FUNCTION_BLOCK "FB_OptEthLink_V1.00"   // FB18, SCL
{ S7_Optimized_Access := 'TRUE' }
VERSION : 0.1
   VAR_INPUT
      IN_xCycleON : Bool;   // Cycle ON
      IN_xCycleONDel : Bool;   // Delayed cycle ON signal
      IN_xGeneralReset : Bool;   // General reset
      IN_xResetAlarms : Bool;   // Reset alarms
      IN_xFaultsEnabled : Bool;   // Faults enabled
      IN_tInterfaceID : Hw_Any;   // Interface ID
      IN_tSmallPckID : Conn_Ouc;   // Connection ID for small packets
      IN_tBigPckID : Conn_Ouc;   // Connection ID for big packets
      IN_uiSmallPckPort : UInt;   // Port small packet
      IN_uiBigPckPort : UInt;   // Port big packet
      IN_rgtStatusYCuts : Array[0.."DMAXYCUTBRIDGE_IND"] of Struct   // Status of YCut
         dDistanceSnapRoll_cmm : DInt;   // Distance from snaproll [mm/100]
         dBridgeStatus : DInt;   // Bridge actual status (1=OutOfProd 3=InProd 4=GlassBreak)
         rgxHeadProdOn : Array[0.."DMAXYHEADS_IND"] of Bool;   // Head#x production status
         rgxFireON : Array[0.."DMAXYHEADS_IND"] of Bool;   // Head#x fire status
         rgxArmON : Array[0.."DMAXYHEADS_IND"] of Bool;   // Head#x arm status
         rgdPosition_cmm : Array[0.."DMAXYHEADS_IND"] of DInt;   // Head#x position [mm/100]
      END_STRUCT;
      IN_rgtStatusXCuts : Array[0.."DMAXXHEADS_IND"] of Struct   // Status of XCuts
         dDistanceFromSnaproll_cmm : DInt;   // Distance from snaproll [mm/100]
         dStatus : DInt;   // XCut actual status (1=Idle 3=Running 7=Faulted)
         dActualCarriagePos_cmm : DInt;   // XCut actual carriage position [mm/100]
         dXCutActualStatus : DInt;   // XCut actual status (1=Disabled 3=Enabled)
         dCutTime_ms : DInt;   // XCut actual cutting time [ms]
      END_STRUCT;
      IN_rgtStatusMarker : Array[0..#DMAXMARKERS_IND] of Struct   // Status of Markers
         dHeadPosition_cmm : DInt;   // Actual head position [mm/100]
         dBridgeProdModeActual : DInt;   // Production modality actual (1=Out of production 3=In production 8=Out of production request 9=In production request)
         dDistanceFromSnaproll_cmm : DInt;   // Distance from snaproll [mm/100]
         dDistanceFromCenterLine_cmm : DInt;   // Distance from center line [mm/100]
         dSpraySpace_cmm : DInt;   // Spray space [mm/100]
         dSpare : DInt;
      END_STRUCT;
   END_VAR
   VAR_IN_OUT
      INO_tInitialize : "GP_OB_Initialize";   // Service bits
      INO_tEncoder : "UDT_Encoder";   // Encoder data
      INO_tOptimizer : "FB_OptManager_V1.00";   // Optimizer manager
      INO_tCaps : "UDT_CapData_Tracking";   // Cap data tracking
      INO_tDefects : "UDT_DefectData_Tracking_Ext";   // Defect data tracking
      INO_tMessage : "UDT_RP_TankMessages";   // Message tank
      INO_tAddMessageFromOpt : "UDT_RP_AddMessageCont_v2";   // Message add for received message
      INO_tAddMessageToOpt : "UDT_RP_AddMessageCont_v2";   // Message add for send message
      INO_xMessageAnomaly : Bool;   // Message anomaly bit
      INO_FB_Markers : "FB_Markers_V1.00";   // Markers FB
   END_VAR
   VAR
      AUX_tStatusPacket : Struct   // Status packet
         dTelID : DInt;   // Telegram identifier
         dTelCount : DInt;   // Telegram counter
         tServiceBit : Struct   // Services bits
            xSpare_24 : Bool;
            xSpare_25 : Bool;
            xSpare_26 : Bool;
            xSpare_27 : Bool;
            xSpare_28 : Bool;
            xSpare_29 : Bool;
            xSpare_30 : Bool;
            xSpare_31 : Bool;
            xSpare_16 : Bool;
            xSpare_17 : Bool;
            xSpare_18 : Bool;
            xSpare_19 : Bool;
            xSpare_20 : Bool;
            xSpare_21 : Bool;
            xSpare_22 : Bool;
            xSpare_23 : Bool;
            xOptRem : Bool;   // Optimizer in remote modality
            xGlassBreak : Bool;   // Glass break
            xSpare_10 : Bool;
            xSpare_11 : Bool;
            xSpare_12 : Bool;
            xSpare_13 : Bool;
            xSpare_14 : Bool;
            xSpare_15 : Bool;
            xSelPCA : Bool;   // Selection PC A
            xSelPCB : Bool;   // Selection PC B
            xSelPLCA : Bool;   // Selection PLC A
            xSelPLCB : Bool;   // Selection PLC B
            xSpare_4 : Bool;
            xSpare_5 : Bool;
            xSpare_6 : Bool;
            xSpare_7 : Bool;
         END_STRUCT;
         dActEnc_cmm : DInt;   // Actual encoder counter [mm/100]
         dActLehrSpeed_mm_min : DInt;   // Actuale lehr speed [mm/min]
         dDecLinePos_cmm : DInt;   // Decision line position [mm/100]
         dLastTargetEnc_cmm : DInt;   // Actual position last plate line [mm/100]
         dLastPlateID : DInt;   // Last plate ID
         dLastPlateLength_cmm : DInt;   // Last plate length [mm/100]
         dLastMapID : DInt;   // Last Map ID
         dSpare3 : DInt;   // Spare
         dRibbonGrossWidth_cmm : DInt;   // Ribbon gross width [mm/100]
         dSpare4 : DInt;   // Spare
         dRibbonNetWidth_cmm : DInt;   // Ribbon net width [mm/100]
         dRibbonWander_cmm : DInt;   // Ribbon wander [mm/100]
         dWanderRecTh_cmm : DInt;   // Ribbon wander recovery threshold [mm/100]
         dLineSpeed_mm_min : DInt;   // Line speed [mm/min]
         dSpare6 : DInt;   // Spare
         dSpare7 : DInt;   // Spare
         dSpare8 : DInt;   // Spare
         dSpare9 : DInt;   // Spare
         dSpare10 : DInt;   // Spare
         dSpare11 : DInt;   // Spare
         dBridgeAStatus : DInt;   // Bridge A status (1=OutOfProd 2=InProd 3=Locked)
         rgdBridgeAHeadxStatus : Array[0..#DMAXYHEADS_IND] of DInt;   // Bridge A headx status (1=OutOfProd 2=InProd 5=Firing)
         rgdBridgeAHeadPos_cmm : Array[0..#DMAXYHEADS_IND] of DInt;   // Bridge A headx position [mm/100]
         dSpare12 : DInt;
         dSpare13 : DInt;
         dSpare14 : DInt;
         dSpare15 : DInt;
         dSpare16 : DInt;
         dBridgeBStatus : DInt;   // Bridge B status (1=OutOfProd 2=InProd 3=Locked)
         rgdBridgeBHeadxStatus : Array[0..#DMAXYHEADS_IND] of DInt;   // Bridge B headx status (1=OutOfProd 2=InProd 5=Firing)
         rgdBridgeBHeadPos_cmm : Array[0..#DMAXYHEADS_IND] of DInt;   // Bridge B headx position [mm/100]
         rgdMarkerState : Array[0..#DMAXMARKERS_IND] of DInt;   // Markers state (1=OutOfProd 3=InProd 7=Anomaly)
         rgdMarkerPos_cmm : Array[0..#DMAXMARKERS_IND] of DInt;   // Markers actual position [mm/100]
         rgdMarkerDistSnap_cmm : Array[0..#DMAXMARKERS_IND] of DInt;   // Markers distance from snaproll [mm/100]
         rgdMarkerSprayTime_ms : Array[0..#DMAXMARKERS_IND] of DInt;   // Markers spray time [ms]
         rgdXCutsState : Array[0..#DMAXXCUT_IND] of DInt;   // XCuts state
         rgdXCutsTimes_ms : Array[0..#DMAXXCUT_IND] of DInt;   // XCuts timing [ms]
         dSpare22 : DInt;
      END_STRUCT;
      AUX_tPlatePacket : Struct   // Plate packet
         dTelID : DInt;   // Telegram identifier
         dTelCounter : DInt;   // Telegram counter
         dPlateHead_cmm : DInt;   // Plate head counter [mm/100]
         rgdLiteID : Array[0..#DMAXLITE_IND] of DInt;   // Lite ID
         rgdProductionID : Array[0..#DMAXLITE_IND] of DInt;   // Production ID
         rgdQualityID : Array[0..#DMAXLITE_IND] of DInt;   // Quality ID
         rgdLiteWidth_cmm : Array[0..#DMAXLITE_IND] of DInt;   // Lite width [mm/100]
         rgdDestMain : Array[0..#DMAXLITE_IND] of LInt;   // Main destination [mask]
         rgdDestAlt : Array[0..#DMAXLITE_IND] of LInt;   // Alternative destination [mask]
         rgdDest2Nd : Array[0..#DMAXLITE_IND] of LInt;   // Second choice destination [mask]
         rgdCulletCause : Array[0..#DMAXLITE_IND] of DInt;   // Cullet cause
         dNumLiteCap : DInt;   // Number of lites in cap
         dCapLength_cmm : DInt;   // Cap length [mm/100]
         dTotCapWidth_cmm : DInt;   // Total cap width [mm/100]
         dColorID : DInt;   // Color ID [mm/100]
         dCapThick_cmm : DInt;   // Cap thickness [mm/100]
         dGeomID : DInt;   // Geometrical ID
         dTrimWidthOper_cmm : DInt;   // Trim width operator side [mm/100]
         dTrimWidthOpOper_cmm : DInt;   // Trim width opposite operator side [mm/100]
         dWanderRec_cmm : DInt;   // Wander recoverd by YCut [mm/100]
         dYBridgeToCut : DInt;   // YCut bridge to cut
         rgxYHeadMask : Array[0..#DMAXYHEADSBITS_IND] of Bool;   // YCut head mask to cut
         rgYBridgePos_cmm : Array[0..#DMAXYHEADS_IND] of DInt;   // YCut head position
         rgxCutMissionHead : Array[0..#DMAXBITSXCUT_INDEX] of Bool;   // XCut mission head
         rgxCutMissionTail : Array[0..#DMAXBITSXCUT_INDEX] of Bool;   // XCut mission tail
         tGeneralFlags : Struct
            xClearCap : Bool;   // Clear cap
            xAutoTrim : Bool;   // Automatic trime selection
            xAutoSnap : Bool;   // Automatic snap bar selection
            xAutoSep : Bool;   // Automatic separator roll selection
            xTripleOpSide : Bool;   // Triple border on operator side
            xTripleOppoOpSide : Bool;   // Triple border on operator opposite side
            xDoubleBorder : Bool;   // Double border enabled
            xYCutSampleTest : Bool;   // YCut sample test
            xIsFixedCap : Bool;   // Is a fixed cap
            xSpare_9 : Bool;
            xSpare_10 : Bool;
            xSpare_11 : Bool;
            xSpare_12 : Bool;
            xSpare_13 : Bool;
            xSpare_14 : Bool;
            xSpare_15 : Bool;
            xSpare_16 : Bool;
            xSpare_17 : Bool;
            xSpare_18 : Bool;
            xSpare_19 : Bool;
            xSpare_20 : Bool;
            xSpare_21 : Bool;
            xSpare_22 : Bool;
            xSpare_23 : Bool;
            xSpare_24 : Bool;
            xSpare_25 : Bool;
            xSpare_26 : Bool;
            xSpare_27 : Bool;
            xSpare_28 : Bool;
            xSpare_29 : Bool;
            xSpare_30 : Bool;
            xSpare_31 : Bool;
         END_STRUCT;
         rgtLiteFlags : Array[0..#DMAXLITE_IND] of Struct
            xPow1Req : Bool;   // Powder #1 request
            xPow2Req : Bool;   // Powder #2 request
            xSatPlate : Bool;   // Saturation plate
            xGeomInsp : Bool;   // Geometrical inspection
            xPrint1 : Bool;   // Print #1 top
            xPrint2 : Bool;   // Print #1 bottom
            xSpare_6 : Bool;
            xSpare_7 : Bool;
            xSpare_8 : Bool;
            xSpare_9 : Bool;
            xSpare_10 : Bool;
            xSpare_11 : Bool;
            xSpare_12 : Bool;
            xSpare_13 : Bool;
            xSpare_14 : Bool;
            xSpare_15 : Bool;
            xMarkHomeHead : Bool;   // Laser mark home head
            xMarkHomeTail : Bool;   // Laser mark home tail
            xMarkCenterHead : Bool;   // Laser mark center head
            xMarkCenterTail : Bool;   // Laser mark center tail
            xMarkFarHead : Bool;   // Laser mark far head
            xMarkFarTail : Bool;   // Laser mark far tail
            xSpare_22 : Bool;
            xSpare_23 : Bool;
            xSpare_24 : Bool;
            xSpare_25 : Bool;
            xSpare_26 : Bool;
            xSpare_27 : Bool;
            xSpare_28 : Bool;
            xSpare_29 : Bool;
            xSpare_30 : Bool;
            xSpare_31 : Bool;   // This lite has a linked cap
         END_STRUCT;
         dExtBordOp : DInt;   // External border operator side
         dIntBordOp : DInt;   // Internal border operator side
         dExtBordOppoOp : DInt;   // External border opposite operator side
         dIntBordOppoOp : DInt;   // Internal border operator side
         rgdBumps : Array[0..#DMAXBUMP_IND] of DInt;   // Bumps splitter
         rgxChevrons : Array[0..#DMAXCHEVRON_IND] of Bool;   // Chevron rolls
         dPlateToPlate_cmm : DInt;   // Plate to plate distance [mm/100]
         dIndexPlateConv : DInt;   // Index plate convoy
         dMaxPlateConv : DInt;   // Max plate convoy
         dConvLength_cmm : DInt;   // Convoy length [mm/100]
         dMinWidth_cmm : DInt;   // Minimum width in production [mm/100]
         dMaxWidth_cmm : DInt;   // Maximum width in production [mm/100]
         dMinLength_cmm : DInt;   // Minimum length in production [mm/100]
         dMaxLength_cmm : DInt;   // Maximum length in production [mm/100]
         dCapID : DInt;   // Cap total ID
         rgdMapPlateID : Array[0..#DMAXLITE_IND] of DInt;   // Map plate ID
         dTripleEdgeOpSide_cmm : DInt;   // Triple edge operator side [mm/100]
         dTripleEdgeOppoOpSide_cmm : DInt;   // Triple edge operator opposite side [mm/100]
         dTripleEdgeHeadOpSide : DInt;   // Triple edge head selection operator side
         dTripleEdgeHeadOppoOpSide : DInt;   // Triple edge head selection oppositio operator side
         dFixedCapProdId : DInt;   // Fixed cap production ID
         rgdSpare : Array[0..10] of DInt;
      END_STRUCT;
      AUX_tDefectPacket : Struct   // Defect packet
         dTelID : DInt;   // Telegram identifier
         dTelCount : DInt;   // Telegram counter
         dNumDefect : DInt;   // Number of defect on packet
         dSpare : DInt;
         dSpare_1 : DInt;
         rgtDefects : Array[0..#DMAXDEFECTS_IND] of Struct
            dID : DInt;   // Defects ID
            dClass : DInt;   // Defects Class
            dSubtype : DInt;   // Defects Subtype
            dPosX_cmm : DInt;   // Defect position X [mm/100]
            dPosY_cmm : DInt;   // Defect position Y [mm/100]
            dTLength_cmm : DInt;   // Total length [mm/100]
            dTWidth_cmm : DInt;   // Total width [mm/100]
            dCLength_cmm : DInt;   // Core length [mm/100]
            dCWidth_cmm : DInt;   // Core width [mm/100]
            dDLength_cmm : DInt;   // Distortion length [mm/100]
            dDWidth_cmm : DInt;   // Distortion width [mm/100]
            dOptDist_mdptr : DInt;   // Optical distortion value [mdptr]
         END_STRUCT;
      END_STRUCT;
      AUX_tMessagePacketToOpt : Struct   // Message packet
         dTelID : DInt;   // Telegram identifier
         dTelCount : DInt;   // Telegram counter
         dNumMessage : DInt;   // Number of message on packet
         dSpare : DInt;
         rgtMessage : Array[0..#DMAXMESSAGEPACKET_IND] of Struct
            dCodeEvent : DInt;
            dEvent1 : DInt;
            dEvent2 : DInt;
            dEvent3 : DInt;
            dEvent4 : DInt;
            dEvent5 : DInt;
            dEvent6 : DInt;
            dEvent7 : DInt;
            dEvent8 : DInt;
            dEvent9 : DInt;
            dEvent10 : DInt;
         END_STRUCT;
      END_STRUCT;
      AUX_tMessagePacketFromOpt : Struct   // Message packet
         dTelID : DInt;   // Telegram identifier
         dTelCount : DInt;   // Telegram counter
         dNumMessage : DInt;   // Number of message on packet
         dSpare : DInt;
         rgtMessage : Array[0..#DMAXMESSAGEPACKET_IND] of Struct
            dCodeEvent : DInt;
            dEvent1 : DInt;
            dEvent2 : DInt;
            dEvent3 : DInt;
            dEvent4 : DInt;
            dEvent5 : DInt;
            dEvent6 : DInt;
            dEvent7 : DInt;
            dEvent8 : DInt;
            dEvent9 : DInt;
            dEvent10 : DInt;
         END_STRUCT;
      END_STRUCT;
      AUX_dNumPlatePacket : DInt;   // Number of plate on buffer
      AUX_rgtPlatePacketArray : Array[0..#DMAXPLATEPACKET_IND] of Struct   // Array buffer of plate
         dTelID : DInt;   // Telegram identifier
         dTelCounter : DInt;   // Telegram counter
         dPlateHead_cmm : DInt;   // Plate head counter [mm/100]
         rgdLiteID : Array[0..#DMAXLITE_IND] of DInt;   // Lite ID
         rgdProductionID : Array[0..#DMAXLITE_IND] of DInt;   // Production ID
         rgdQualityID : Array[0..#DMAXLITE_IND] of DInt;   // Quality ID
         rgdLiteWidth_cmm : Array[0..#DMAXLITE_IND] of DInt;   // Lite width [mm/100]
         rgdDestMain : Array[0..#DMAXLITE_IND] of LInt;   // Main destination [mask]
         rgdDestAlt : Array[0..#DMAXLITE_IND] of LInt;   // Alternative destination [mask]
         rgdDest2Nd : Array[0..#DMAXLITE_IND] of LInt;   // Second choice destination [mask]
         rgdCulletCause : Array[0..#DMAXLITE_IND] of DInt;   // Cullet cause
         dNumLiteCap : DInt;   // Number of lites in cap
         dCapLength_cmm : DInt;   // Cap length [mm/100]
         dTotCapWidth_cmm : DInt;   // Total cap width [mm/100]
         dColorID : DInt;   // Color ID [mm/100]
         dCapThick_cmm : DInt;   // Cap thickness [mm/100]
         dGeomID : DInt;   // Geometrical ID
         dTrimWidthOper_cmm : DInt;   // Trim width operator side [mm/100]
         dTrimWidthOpOper_cmm : DInt;   // Trim width opposite operator side [mm/100]
         dWanderRec_cmm : DInt;   // Wander recoverd by YCut [mm/100]
         dYBridgeToCut : DInt;   // YCut bridge to cut
         rgxYHeadMask : Array[0..#DMAXYHEADSBITS_IND] of Bool;   // YCut head mask to cut
         rgYBridgePos_cmm : Array[0..#DMAXYHEADS_IND] of DInt;   // YCut head position
         rgxCutMissionHead : Array[0..#DMAXBITSXCUT_INDEX] of Bool;   // XCut mission head
         rgxCutMissionTail : Array[0..#DMAXBITSXCUT_INDEX] of Bool;   // XCut mission tail
         tGeneralFlags : Struct
            xClearCap : Bool;   // Clear cap
            xAutoTrim : Bool;   // Automatic trime selection
            xAutoSnap : Bool;   // Automatic snap bar selection
            xAutoSep : Bool;   // Automatic separator roll selection
            xTripleOpSide : Bool;   // Triple border on operator side
            xTripleOppoOpSide : Bool;   // Triple border on operator opposite side
            xDoubleBorder : Bool;   // Double border enabled
            xYCutSampleTest : Bool;   // YCut sample test
            xIsFixedCap : Bool;   // Is a fixed cap
            xSpare_9 : Bool;
            xSpare_10 : Bool;
            xSpare_11 : Bool;
            xSpare_12 : Bool;
            xSpare_13 : Bool;
            xSpare_14 : Bool;
            xSpare_15 : Bool;
            xSpare_16 : Bool;
            xSpare_17 : Bool;
            xSpare_18 : Bool;
            xSpare_19 : Bool;
            xSpare_20 : Bool;
            xSpare_21 : Bool;
            xSpare_22 : Bool;
            xSpare_23 : Bool;
            xSpare_24 : Bool;
            xSpare_25 : Bool;
            xSpare_26 : Bool;
            xSpare_27 : Bool;
            xSpare_28 : Bool;
            xSpare_29 : Bool;
            xSpare_30 : Bool;
            xSpare_31 : Bool;
         END_STRUCT;
         rgtLiteFlags : Array[0..#DMAXLITE_IND] of Struct
            xPow1Req : Bool;   // Powder #1 request
            xPow2Req : Bool;   // Powder #2 request
            xSatPlate : Bool;   // Saturation plate
            xGeomInsp : Bool;   // Geometrical inspection
            xPrint1 : Bool;   // Print #1 top
            xPrint2 : Bool;   // Print #1 bottom
            xSpare_6 : Bool;
            xSpare_7 : Bool;
            xSpare_8 : Bool;
            xSpare_9 : Bool;
            xSpare_10 : Bool;
            xSpare_11 : Bool;
            xSpare_12 : Bool;
            xSpare_13 : Bool;
            xSpare_14 : Bool;
            xSpare_15 : Bool;
            xMarkHomeHead : Bool;   // Laser mark home head
            xMarkHomeTail : Bool;   // Laser mark home tail
            xMarkCenterHead : Bool;   // Laser mark center head
            xMarkCenterTail : Bool;   // Laser mark center tail
            xMarkFarHead : Bool;   // Laser mark far head
            xMarkFarTail : Bool;   // Laser mark far tail
            xSpare_22 : Bool;
            xSpare_23 : Bool;
            xSpare_24 : Bool;
            xSpare_25 : Bool;
            xSpare_26 : Bool;
            xSpare_27 : Bool;
            xSpare_28 : Bool;
            xSpare_29 : Bool;
            xSpare_30 : Bool;
            xSpare_31 : Bool;   // This lite has a linked cap
         END_STRUCT;
         dExtBordOp : DInt;   // External border operator side
         dIntBordOp : DInt;   // Internal border operator side
         dExtBordOppoOp : DInt;   // External border opposite operator side
         dIntBordOppoOp : DInt;   // Internal border operator side
         rgdBumps : Array[0..#DMAXBUMP_IND] of DInt;   // Bumps splitter
         rgxChevrons : Array[0..#DMAXCHEVRON_IND] of Bool;   // Chevron rolls
         dPlateToPlate_cmm : DInt;   // Plate to plate distance [mm/100]
         dIndexPlateConv : DInt;   // Index plate convoy
         dMaxPlateConv : DInt;   // Max plate convoy
         dConvLength_cmm : DInt;   // Convoy length [mm/100]
         dMinWidth_cmm : DInt;   // Minimum width in production [mm/100]
         dMaxWidth_cmm : DInt;   // Maximum width in production [mm/100]
         dMinLength_cmm : DInt;   // Minimum length in production [mm/100]
         dMaxLength_cmm : DInt;   // Maximum length in production [mm/100]
         dCapID : DInt;   // Cap total ID
         rgdMapPlateID : Array[0..#DMAXLITE_IND] of DInt;   // Map plate ID
         dTripleEdgeOpSide_cmm : DInt;   // Triple edge operator side [mm/100]
         dTripleEdgeOppoOpSide_cmm : DInt;   // Triple edge operator opposite side [mm/100]
         dTripleEdgeHeadOpSide : DInt;   // Triple edge head selection operator side
         dTripleEdgeHeadOppoOpSide : DInt;   // Triple edge head selection oppositio operator side
         dFixedCapProdId : DInt;   // Fixed cap production ID
         rgdSpare : Array[0..10] of DInt;
      END_STRUCT;
      AUX_rgb500SendBytePck : Array[0..#DSMALLSIZEPACKET_IND] of Byte;   // Byte array small size packet
      AUX_rgb500RecvBytePck : Array[0..#DSMALLSIZEPACKET_IND] of Byte;   // Byte array small size packet
      AUX_rgb1000SendBytePck : Array[0..#DBIGSIZEPACKET_IND] of Byte;   // Byte array big size packet
      AUX_rgb1000RecvBytePck : Array[0..#DBIGSIZEPACKET_IND] of Byte;   // Byte array big size packet
      FB_TSendSmall : TSEND_C;   // FB send small
      FB_TRecvSmall : TRCV_C;   // FB receive small
      FB_TSendBig : TSEND_C;   // FB send big
      FB_TRecvBig : TRCV_C;   // FB receive big
      AUX_tConnDataSmall : TCON_IP_v4;   // Connection small data structure
      AUX_tConnDataBig : TCON_IP_v4;   // Connection big data structure
      tPhasesNetworkSmall : Struct   // Phases network small
         xSendBuffer : Bool;   // Send buffer in progress
         xEndSendBuffer : Bool;   // End send buffer in progress
         xSpare2 : Bool;
         xSpare3 : Bool;
         xSpare4 : Bool;
         xSpare5 : Bool;
         xSpare6 : Bool;
         xSpare7 : Bool;
         xSpare8 : Bool;
         xSpare9 : Bool;
         xSpare10 : Bool;
         xSpare11 : Bool;
         xSpare12 : Bool;
         xSpare13 : Bool;
         xSpare14 : Bool;
         xSpare15 : Bool;
         xSpare16 : Bool;
         xSpare17 : Bool;
         xSpare18 : Bool;
         xSpare19 : Bool;
         xSpare20 : Bool;
         xSpare21 : Bool;
         xSpare22 : Bool;
         xSpare23 : Bool;
         xSpare24 : Bool;
         xSpare25 : Bool;
         xSpare26 : Bool;
         xSpare27 : Bool;
         xSpare28 : Bool;
         xSpare29 : Bool;
         xSpare30 : Bool;
         xSpare31 : Bool;
      END_STRUCT;
      tPhasesNetworkBig : Struct   // Phases network big
         xSendBuffer : Bool;   // Send buffer in progress
         xEndSendBuffer : Bool;   // End send buffer in progress
         xSpare2 : Bool;
         xSpare3 : Bool;
         xSpare4 : Bool;
         xSpare5 : Bool;
         xSpare6 : Bool;
         xSpare7 : Bool;
         xSpare8 : Bool;
         xSpare9 : Bool;
         xSpare10 : Bool;
         xSpare11 : Bool;
         xSpare12 : Bool;
         xSpare13 : Bool;
         xSpare14 : Bool;
         xSpare15 : Bool;
         xSpare16 : Bool;
         xSpare17 : Bool;
         xSpare18 : Bool;
         xSpare19 : Bool;
         xSpare20 : Bool;
         xSpare21 : Bool;
         xSpare22 : Bool;
         xSpare23 : Bool;
         xSpare24 : Bool;
         xSpare25 : Bool;
         xSpare26 : Bool;
         xSpare27 : Bool;
         xSpare28 : Bool;
         xSpare29 : Bool;
         xSpare30 : Bool;
         xSpare31 : Bool;
      END_STRUCT;
      AUX_xResetSendConnection : Bool;   // Reset send connection
      ST_xRetrySendTelegramSmall : Bool;   // Retry send telegram small
      ST_xRetrySendTelegramBig : Bool;   // Retry send telegram big
      ST_xStatusTelegramAvail : Bool;   // Status telegram available to send
      ST_xDefectTelegramAvail : Bool;   // Defect telegram available to send
      ST_xMessageTelegramAvail : Bool;   // Message telegram available to send
      ST_xSmallChannelConnected : Bool;   // Small channel connected
      ST_xBigChannelConnected : Bool;   // Big channel connected
      AUX_dWaitingNextStatus_ms : DInt;   // Waiting time for next status packet [ms]
   END_VAR
   VAR RETAIN
      AUX_dStatusTelegramCounter : DInt := 1;   // Status telegram counter
      AUX_dDefectTelegramCounter : DInt := 1;   // Defect telegram counter
      AUX_dMessageTelegramCounter : DInt := 1;   // Telegram message counter
   END_VAR
   VAR
      AUX_tEmptyMessage : "UDT_RP_Message_v2";   // Empty message
      tALM : Struct   // HMI Alarms
         tS : Struct   // Stopping faults
            xCh1NotCon : Bool;   // Channel 1 not connected {X|X|X|X|O}
            xCh2NotCon : Bool;   // Channel 2 not connected {X|X|X|X|O}
            xSpare_2 : Bool;
            xSpare_3 : Bool;
            xSpare_4 : Bool;
            xSpare_5 : Bool;
            xSpare_6 : Bool;
            xSpare_7 : Bool;
            xSpare_8 : Bool;
            xSpare_9 : Bool;
            xSpare_10 : Bool;
            xSpare_11 : Bool;
            xSpare_12 : Bool;
            xSpare_13 : Bool;
            xSpare_14 : Bool;
            xSpare_15 : Bool;
            xSpare_16 : Bool;
            xSpare_17 : Bool;
            xSpare_18 : Bool;
            xSpare_19 : Bool;
            xSpare_20 : Bool;
            xSpare_21 : Bool;
            xSpare_22 : Bool;
            xSpare_23 : Bool;
            xSpare_24 : Bool;
            xSpare_25 : Bool;
            xSpare_26 : Bool;
            xSpare_27 : Bool;
            xSpare_28 : Bool;
            xSpare_29 : Bool;
            xSpare_30 : Bool;
            xSpare_31 : Bool;
         END_STRUCT;
         tF : Struct   // Faults
            xSpare_0 : Bool;
            xSpare_1 : Bool;
            xSpare_2 : Bool;
            xSpare_3 : Bool;
            xSpare_4 : Bool;
            xSpare_5 : Bool;
            xSpare_6 : Bool;
            xSpare_7 : Bool;
            xSpare_8 : Bool;
            xSpare_9 : Bool;
            xSpare_10 : Bool;
            xSpare_11 : Bool;
            xSpare_12 : Bool;
            xSpare_13 : Bool;
            xSpare_14 : Bool;
            xSpare_15 : Bool;
            xSpare_16 : Bool;
            xSpare_17 : Bool;
            xSpare_18 : Bool;
            xSpare_19 : Bool;
            xSpare_20 : Bool;
            xSpare_21 : Bool;
            xSpare_22 : Bool;
            xSpare_23 : Bool;
            xSpare_24 : Bool;
            xSpare_25 : Bool;
            xSpare_26 : Bool;
            xSpare_27 : Bool;
            xSpare_28 : Bool;
            xSpare_29 : Bool;
            xSpare_30 : Bool;
            xSpare_31 : Bool;
         END_STRUCT;
         tW : Struct   // Warnings
            xSpare_0 : Bool;
            xSpare_1 : Bool;
            xSpare_2 : Bool;
            xSpare_3 : Bool;
            xSpare_4 : Bool;
            xSpare_5 : Bool;
            xSpare_6 : Bool;
            xSpare_7 : Bool;
            xSpare_8 : Bool;
            xSpare_9 : Bool;
            xSpare_10 : Bool;
            xSpare_11 : Bool;
            xSpare_12 : Bool;
            xSpare_13 : Bool;
            xSpare_14 : Bool;
            xSpare_15 : Bool;
            xSpare_16 : Bool;
            xSpare_17 : Bool;
            xSpare_18 : Bool;
            xSpare_19 : Bool;
            xSpare_20 : Bool;
            xSpare_21 : Bool;
            xSpare_22 : Bool;
            xSpare_23 : Bool;
            xSpare_24 : Bool;
            xSpare_25 : Bool;
            xSpare_26 : Bool;
            xSpare_27 : Bool;
            xSpare_28 : Bool;
            xSpare_29 : Bool;
            xSpare_30 : Bool;
            xSpare_31 : Bool;
         END_STRUCT;
      END_STRUCT;
   END_VAR
   VAR_TEMP
      TMP_dIndex : DInt;
      TMP_dSerializePos : DInt;   // Serialize temporary position
      TMP_iReturn : Int;
      TMP_dValue : DInt;
      TMP_dwMask : DWord;
      TMP_wMask : Word;
      TMP_dCounter : DInt;
      TMP_dRemaining : DInt;
      TMP_rgbDInt : Array[0..3] of Byte;
      TMP_iRetVal : Int;
      TMP_tNewMisMark : "UDT_Marker_Mission_Data";
      TMP_xCallAddTank : Bool;
      TMP_dwValue : DWord;
   END_VAR
   VAR CONSTANT
      DMAXYHEADS : DInt := 16;   // Maximum number of heads
      DMAXYHEADS_IND : DInt := 15;   // Maximum number of heads index (Always -1)
      DMAXYHEADSBITS : DInt := 32;   // Maximum number of heads bits
      DMAXYHEADSBITS_IND : DInt := 31;   // Maximum number of heads bits index (Always -1)
      DMAXMARKERS : DInt := 5;   // Maximum number of markers bridge
      DMAXMARKERS_IND : DInt := 4;   // Maximum number of markers bridge index (Always -1)
      DMAXXCUT : DInt := 5;   // Maximum number of cross cut bridge
      DMAXXCUT_IND : DInt := 4;   // Maximum number of cross cut bridge index (Always -1)
      DMAXLITE : DInt := 12;   // Maximum number of lite
      DMAXLITE_IND : DInt := 11;   // Maximum numer of lite index (Always -1)
      DMAXBITSXCUT : DInt := 32;   // Maximum number of request bits xcuts
      DMAXBITSXCUT_INDEX : DInt := 31;   // Maximum number of request bits xcuts index (Always -1)
      DMAXBUMP : DInt := 12;   // Maximum number of bump
      DMAXBUMP_IND : DInt := 11;   // Maximum numer of bump index (Always -1)
      DMAXCHEVRON : DInt := 32;   // Maximum number of chevron rolls
      DMAXCHEVRON_IND : DInt := 31;   // Maximum number of chevron rolls index (Always -1)
      BCONNTYPE : Byte := 16#0B;   // Optimizer connection type
      DSMALLSIZEPACKET : DInt := 500;   // Size of the small size packet
      DSMALLSIZEPACKET_IND : DInt := 499;   // Size of the small size packet index (Always -1)
      DBIGSIZEPACKET : DInt := 1000;   // Size of the big size packet
      DBIGSIZEPACKET_IND : DInt := 999;   // Size of the big size packet index (Always -1)
      DDELAYSTATUSPACKET_MS : DInt := 500;   // Status packet delay [ms]
      DSTATUSPACKETIDENT : DInt := 16#11111111;   // Status packet identifier
      DDEFECTPACKTIDENT : DInt := 16#22222222;   // Defect packet identifier
      DMESSAGEPACKETIDENT : DInt := 16#33333333;   // Message packet identifier
      DPLATEPACKTIDENT : DInt := 16#44444444;   // Plate packet identifier
      DMESSAGERECVPACKETIDENT : DInt := 16#55555555;   // Message received packet identifier
      DMAXTELEGRAMCOUNTER : DInt := 2000000000;   // Maximum telegram counter
      DMAXDEFECTS : DInt := 10;   // Maximum number of defects
      DMAXDEFECTS_IND : DInt := 9;   // Maximum number of defects index (Always -1)
      DMAXPLATEPACKET : DInt := 5;   // Number maximum of plate packet
      DMAXPLATEPACKET_IND : DInt := 4;   // Number maximum of plate packet index (Always -1)
      DMAXMESSAGEPACKET : DInt := 11;   // Number maximum of message packet
      DMAXMESSAGEPACKET_IND : DInt := 10;   // Number maximum of message packet index (Always -1)
   END_VAR
BEGIN
   IF #IN_xResetAlarms THEN

       #TMP_dwValue := 0;

       SCATTER(IN := #TMP_dwValue,
               OUT => #tALM.tS);

       SCATTER(IN := #TMP_dwValue,
               OUT => #tALM.tF);

       SCATTER(IN := #TMP_dwValue,
               OUT => #tALM.tW);


   END_IF;

   #ST_xSmallChannelConnected := TRUE;
   #ST_xBigChannelConnected := TRUE;

   IF #FB_TSendSmall.s_TDIAG_Status.State <> b#16#04(* OR #FB_TRecvSmall.s_TDIAG_Status.State <> b#16#04*) THEN

       #ST_xRetrySendTelegramSmall := FALSE;
       #ST_xStatusTelegramAvail := FALSE;
       #ST_xMessageTelegramAvail := FALSE;

       #tPhasesNetworkSmall.xSendBuffer := FALSE;
       #tPhasesNetworkSmall.xEndSendBuffer := FALSE;

       #ST_xSmallChannelConnected := FALSE;

       #INO_tDefects.xOptimizerRequireAllDef := TRUE;
   END_IF;

   IF #FB_TRecvBig.s_TRCV.ERROR  THEN
       #ST_xBigChannelConnected := FALSE;
   END_IF;

   //Calculate anomalies
   #tALM.tS.xCh1NotCon := NOT #ST_xSmallChannelConnected;
   #tALM.tS.xCh2NotCon := NOT #ST_xBigChannelConnected;


   IF #IN_xGeneralReset THEN
       #AUX_tConnDataSmall.InterfaceId := #IN_tInterfaceID;
       #AUX_tConnDataSmall.ID := #IN_tSmallPckID;
       #AUX_tConnDataSmall.ConnectionType := #BCONNTYPE;
       #AUX_tConnDataSmall.ActiveEstablished := FALSE;
       #AUX_tConnDataSmall.RemotePort := 0;
       #AUX_tConnDataSmall.LocalPort := #IN_uiSmallPckPort;

       #AUX_tConnDataBig.InterfaceId := #IN_tInterfaceID;
       #AUX_tConnDataBig.ID := #IN_tBigPckID;
       #AUX_tConnDataBig.ConnectionType := #BCONNTYPE;
       #AUX_tConnDataBig.ActiveEstablished := FALSE;
       #AUX_tConnDataBig.RemotePort := 0;
       #AUX_tConnDataBig.LocalPort := #IN_uiBigPckPort;
   END_IF;

   #AUX_dWaitingNextStatus_ms-= #INO_tInitialize.OUT_dExecutionTime_ms;

   IF #AUX_dWaitingNextStatus_ms < 0 THEN
       #AUX_dWaitingNextStatus_ms := 0;
   END_IF;


   IF NOT #ST_xMessageTelegramAvail AND #ST_xSmallChannelConnected THEN

       IF #INO_tMessage.dNumberOfMessage > 0 THEN
           #AUX_tMessagePacketToOpt.dTelID := #DMESSAGEPACKETIDENT;
           #AUX_tMessagePacketToOpt.dTelCount := #AUX_dMessageTelegramCounter;

           #TMP_dCounter := 0;

           WHILE (#TMP_dCounter < #DMAXMESSAGEPACKET) AND (#TMP_dCounter < #INO_tMessage.dNumberOfMessage) DO

               #AUX_tMessagePacketToOpt.rgtMessage[#TMP_dCounter].dCodeEvent := #INO_tMessage.rgtMessages[#TMP_dCounter].dCodeEvent;
               #AUX_tMessagePacketToOpt.rgtMessage[#TMP_dCounter].dEvent1 := #INO_tMessage.rgtMessages[#TMP_dCounter].dEvent1;
               #AUX_tMessagePacketToOpt.rgtMessage[#TMP_dCounter].dEvent2 := #INO_tMessage.rgtMessages[#TMP_dCounter].dEvent2;
               #AUX_tMessagePacketToOpt.rgtMessage[#TMP_dCounter].dEvent3 := #INO_tMessage.rgtMessages[#TMP_dCounter].dEvent3;
               #AUX_tMessagePacketToOpt.rgtMessage[#TMP_dCounter].dEvent4 := #INO_tMessage.rgtMessages[#TMP_dCounter].dEvent4;
               #AUX_tMessagePacketToOpt.rgtMessage[#TMP_dCounter].dEvent5 := #INO_tMessage.rgtMessages[#TMP_dCounter].dEvent5;
               #AUX_tMessagePacketToOpt.rgtMessage[#TMP_dCounter].dEvent6 := #INO_tMessage.rgtMessages[#TMP_dCounter].dEvent6;
               #AUX_tMessagePacketToOpt.rgtMessage[#TMP_dCounter].dEvent7 := #INO_tMessage.rgtMessages[#TMP_dCounter].dEvent7;
               #AUX_tMessagePacketToOpt.rgtMessage[#TMP_dCounter].dEvent8 := #INO_tMessage.rgtMessages[#TMP_dCounter].dEvent8;
               #AUX_tMessagePacketToOpt.rgtMessage[#TMP_dCounter].dEvent9 := #INO_tMessage.rgtMessages[#TMP_dCounter].dEvent9;
               #AUX_tMessagePacketToOpt.rgtMessage[#TMP_dCounter].dEvent10 := #INO_tMessage.rgtMessages[#TMP_dCounter].dEvent10;

               #INO_tMessage.rgtMessages[#TMP_dCounter] := #AUX_tEmptyMessage;

               #TMP_dCounter += 1;

           END_WHILE;

           //Clear the remaining packet
           FOR #TMP_dIndex := #TMP_dCounter TO #DMAXMESSAGEPACKET - 1 DO
               #AUX_tMessagePacketToOpt.rgtMessage[#TMP_dIndex].dCodeEvent := 0;
               #AUX_tMessagePacketToOpt.rgtMessage[#TMP_dIndex].dEvent1 := 0;
               #AUX_tMessagePacketToOpt.rgtMessage[#TMP_dIndex].dEvent2 := 0;
               #AUX_tMessagePacketToOpt.rgtMessage[#TMP_dIndex].dEvent3 := 0;
               #AUX_tMessagePacketToOpt.rgtMessage[#TMP_dIndex].dEvent4 := 0;
               #AUX_tMessagePacketToOpt.rgtMessage[#TMP_dIndex].dEvent5 := 0;
               #AUX_tMessagePacketToOpt.rgtMessage[#TMP_dIndex].dEvent6 := 0;
               #AUX_tMessagePacketToOpt.rgtMessage[#TMP_dIndex].dEvent7 := 0;
               #AUX_tMessagePacketToOpt.rgtMessage[#TMP_dIndex].dEvent8 := 0;
               #AUX_tMessagePacketToOpt.rgtMessage[#TMP_dIndex].dEvent9 := 0;
               #AUX_tMessagePacketToOpt.rgtMessage[#TMP_dIndex].dEvent10 := 0;
           END_FOR;

           #AUX_tMessagePacketToOpt.dNumMessage := #TMP_dCounter;
           #AUX_dMessageTelegramCounter+= 1;
           #ST_xMessageTelegramAvail := TRUE;
           #TMP_dRemaining := #INO_tMessage.dNumberOfMessage - #TMP_dCounter;

           IF #TMP_dRemaining > 0 THEN
               #TMP_iRetVal :=  MOVE_BLK_VARIANT(   SRC:= #INO_tMessage.rgtMessages, 
                                   COUNT:=DINT_TO_UDINT(#TMP_dRemaining), 
                                   SRC_INDEX:=#TMP_dCounter, 
                                   DEST_INDEX:=0, 
                                   DEST=>#INO_tMessage.rgtMessages);
               //Reset the remaining
               FOR #TMP_dIndex := #TMP_dRemaining TO #INO_tMessage.dNumberOfMessage - 1 DO
                   #INO_tMessage.rgtMessages[#TMP_dIndex] := #AUX_tEmptyMessage;
               END_FOR;

               #INO_tMessage.dNumberOfMessage := #TMP_dRemaining;

           ELSE
               #INO_tMessage.dNumberOfMessage := 0;
           END_IF;
       END_IF;
   END_IF;

   //Prepare defect telegram
   IF NOT #ST_xDefectTelegramAvail AND #ST_xSmallChannelConnected  THEN

       IF #INO_tDefects.tDefectsForOpt.dNumberOfDefect > 0 THEN

           #AUX_tDefectPacket.dTelID := #DDEFECTPACKTIDENT;
           #AUX_tDefectPacket.dTelCount := #AUX_dDefectTelegramCounter;
           #AUX_tDefectPacket.dNumDefect := #INO_tDefects.tDefectsForOpt.dNumberOfDefect;

           FOR #TMP_dIndex := 0 TO #DMAXDEFECTS_IND DO

               #AUX_tDefectPacket.rgtDefects[#TMP_dIndex].dID := #INO_tDefects.tDefectsForOpt.rgtDefects[#TMP_dIndex].dID;
               #AUX_tDefectPacket.rgtDefects[#TMP_dIndex].dClass := #INO_tDefects.tDefectsForOpt.rgtDefects[#TMP_dIndex].dClass;
               #AUX_tDefectPacket.rgtDefects[#TMP_dIndex].dSubtype := #INO_tDefects.tDefectsForOpt.rgtDefects[#TMP_dIndex].dSubType;
               #AUX_tDefectPacket.rgtDefects[#TMP_dIndex].dPosX_cmm := #INO_tDefects.tDefectsForOpt.rgtDefects[#TMP_dIndex].dXPosition_cmm;
               #AUX_tDefectPacket.rgtDefects[#TMP_dIndex].dPosY_cmm := #INO_tDefects.tDefectsForOpt.rgtDefects[#TMP_dIndex].dYPosition_cmm;
               #AUX_tDefectPacket.rgtDefects[#TMP_dIndex].dCLength_cmm := #INO_tDefects.tDefectsForOpt.rgtDefects[#TMP_dIndex].dCoreLength_um;
               #AUX_tDefectPacket.rgtDefects[#TMP_dIndex].dCWidth_cmm := #INO_tDefects.tDefectsForOpt.rgtDefects[#TMP_dIndex].dCoreWidth_um;
               #AUX_tDefectPacket.rgtDefects[#TMP_dIndex].dDLength_cmm := #INO_tDefects.tDefectsForOpt.rgtDefects[#TMP_dIndex].dDistLength_um;
               #AUX_tDefectPacket.rgtDefects[#TMP_dIndex].dDWidth_cmm := #INO_tDefects.tDefectsForOpt.rgtDefects[#TMP_dIndex].dDistWidth_um;
               #AUX_tDefectPacket.rgtDefects[#TMP_dIndex].dTLength_cmm := #INO_tDefects.tDefectsForOpt.rgtDefects[#TMP_dIndex].dTotalLength_um;
               #AUX_tDefectPacket.rgtDefects[#TMP_dIndex].dTWidth_cmm := #INO_tDefects.tDefectsForOpt.rgtDefects[#TMP_dIndex].dTotalWidth_um;
               #AUX_tDefectPacket.rgtDefects[#TMP_dIndex].dOptDist_mdptr := #INO_tDefects.tDefectsForOpt.rgtDefects[#TMP_dIndex].dOptValue_mdptr;

           END_FOR;

           #ST_xDefectTelegramAvail := TRUE;
           #AUX_dDefectTelegramCounter += 1;
           #INO_tDefects.tDefectsForOpt.dNumberOfDefect := 0;
       END_IF;

   END_IF;

   //Prepare status telegram
   IF NOT #ST_xStatusTelegramAvail AND #AUX_dWaitingNextStatus_ms = 0 AND #ST_xSmallChannelConnected THEN

       #AUX_dWaitingNextStatus_ms := #DDELAYSTATUSPACKET_MS;

       //Prepare data
       #AUX_tStatusPacket.dTelID :=  #DSTATUSPACKETIDENT;
       #AUX_tStatusPacket.dSpare22 := #DSTATUSPACKETIDENT;
       #AUX_tStatusPacket.dTelCount := #AUX_dStatusTelegramCounter;


       IF "FB_OptManager_V1_00_IDB".tHMR.dSelOptimizer = 1 THEN
           #AUX_tStatusPacket.tServiceBit.xSelPCA := TRUE;
           #AUX_tStatusPacket.tServiceBit.xSelPCB := FALSE;
       ELSE
           #AUX_tStatusPacket.tServiceBit.xSelPCA := FALSE;
           #AUX_tStatusPacket.tServiceBit.xSelPCB := TRUE;
       END_IF;

       #AUX_tStatusPacket.tServiceBit.xSelPLCA := TRUE;
       #AUX_tStatusPacket.tServiceBit.xSelPLCB := FALSE;
       #AUX_tStatusPacket.tServiceBit.xOptRem := TRUE;
       #AUX_tStatusPacket.tServiceBit.xGlassBreak := FALSE;

       #AUX_tStatusPacket.dActEnc_cmm := #INO_tEncoder.dActualEncoderCounter_cmm;
       #AUX_tStatusPacket.dActLehrSpeed_mm_min := #INO_tEncoder.dActSpeedValue_mm_min;
       #AUX_tStatusPacket.dDecLinePos_cmm := #INO_tOptimizer.tHMR.dDecisionLinePosition_cmm;
       #AUX_tStatusPacket.dLastTargetEnc_cmm := #INO_tCaps.dLastTargetLineValue_cmm;
       #AUX_tStatusPacket.dLastPlateID := #INO_tCaps.dLastValidCapID;

       #AUX_tStatusPacket.dRibbonGrossWidth_cmm := #INO_tOptimizer.tHMR.rgtRibbonData[#INO_tOptimizer.tHMW.dSelectRibbonDataSource].dGrossWidth_cmm;
       #AUX_tStatusPacket.dRibbonNetWidth_cmm := #INO_tOptimizer.tHMR.rgtRibbonData[#INO_tOptimizer.tHMW.dSelectRibbonDataSource].dNetWidth_cmm;

       #AUX_tStatusPacket.dWanderRecTh_cmm := #INO_tOptimizer.tHMW.dWanderRecThr_cmm;

       IF #INO_tOptimizer.tHMW.dSelectWanderMode = 0 THEN
           #AUX_tStatusPacket.dRibbonWander_cmm := #INO_tOptimizer.tHMR.rgtRibbonData[#INO_tOptimizer.tHMW.dSelectWanderDataSource].dNetWander_cmm + #INO_tOptimizer.tHMW.dWanderOffset_cmm;
       ELSE
           #AUX_tStatusPacket.dRibbonWander_cmm := #INO_tOptimizer.tHMR.rgtRibbonData[#INO_tOptimizer.tHMW.dSelectWanderDataSource].dGrossWander_cmm + #INO_tOptimizer.tHMW.dWanderOffset_cmm;
       END_IF;


       CASE #IN_rgtStatusYCuts[0].dBridgeStatus OF

           1:
               #AUX_tStatusPacket.dBridgeAStatus := 1;//Out of production
           3: #AUX_tStatusPacket.dBridgeAStatus := 2;
           4: #AUX_tStatusPacket.dBridgeAStatus := 2; //Glass break, out of production for optimizer

       END_CASE;

       CASE #IN_rgtStatusYCuts[1].dBridgeStatus OF

           1:
               #AUX_tStatusPacket.dBridgeBStatus := 1;//Out of production
           3: #AUX_tStatusPacket.dBridgeBStatus := 2;
           4: #AUX_tStatusPacket.dBridgeBStatus := 2; //Glass break, out of production for optimizer

       END_CASE;

       FOR #TMP_dIndex := 0 TO #DMAXYHEADS_IND DO

           IF #IN_rgtStatusYCuts[0].rgxHeadProdOn[#TMP_dIndex] = TRUE THEN
               #AUX_tStatusPacket.rgdBridgeAHeadxStatus[#TMP_dIndex] := 2;
           ELSE
               #AUX_tStatusPacket.rgdBridgeAHeadxStatus[#TMP_dIndex] := 1;
           END_IF;

           IF #IN_rgtStatusYCuts[1].rgxHeadProdOn[#TMP_dIndex] = TRUE THEN
               #AUX_tStatusPacket.rgdBridgeBHeadxStatus[#TMP_dIndex] := 2;
           ELSE
               #AUX_tStatusPacket.rgdBridgeBHeadxStatus[#TMP_dIndex] := 1;
           END_IF;

       END_FOR;

       #AUX_tStatusPacket.rgdBridgeAHeadPos_cmm := #IN_rgtStatusYCuts[0].rgdPosition_cmm;
       #AUX_tStatusPacket.rgdBridgeBHeadPos_cmm := #IN_rgtStatusYCuts[1].rgdPosition_cmm;

       FOR #TMP_dIndex := 0 TO #DMAXMARKERS_IND DO

           #AUX_tStatusPacket.rgdMarkerDistSnap_cmm[#TMP_dIndex] := #IN_rgtStatusMarker[#TMP_dIndex].dDistanceFromSnaproll_cmm;
           #AUX_tStatusPacket.rgdMarkerPos_cmm[#TMP_dIndex] := #IN_rgtStatusMarker[#TMP_dIndex].dHeadPosition_cmm;
           #AUX_tStatusPacket.rgdMarkerSprayTime_ms[#TMP_dIndex] := REAL_TO_DINT(DINT_TO_REAL(#IN_rgtStatusMarker[#TMP_dIndex].dSpraySpace_cmm) / #INO_tEncoder.rActSpeedValue_cmm_ms);

           CASE #IN_rgtStatusMarker[#TMP_dIndex].dBridgeProdModeActual OF

               1: #AUX_tStatusPacket.rgdMarkerState[#TMP_dIndex] := 1;//Out of production
               3: #AUX_tStatusPacket.rgdMarkerState[#TMP_dIndex] := 2;//In production
               8: #AUX_tStatusPacket.rgdMarkerState[#TMP_dIndex] := 1;//Out of production
               9: #AUX_tStatusPacket.rgdMarkerState[#TMP_dIndex] := 1;//Out of production

           END_CASE;

       END_FOR; 

       FOR #TMP_dIndex := 0 TO "DMAXXHEADS_IND" DO

           CASE #IN_rgtStatusXCuts[#TMP_dIndex].dXCutActualStatus OF

               1: #AUX_tStatusPacket.rgdXCutsState[#TMP_dIndex] := 0;
               3: #AUX_tStatusPacket.rgdXCutsState[#TMP_dIndex] := 1;

           END_CASE;

           #AUX_tStatusPacket.rgdXCutsTimes_ms[#TMP_dIndex] := #IN_rgtStatusXCuts[#TMP_dIndex].dCutTime_ms;

       END_FOR;

       IF #AUX_dStatusTelegramCounter >= #DMAXTELEGRAMCOUNTER THEN
           #AUX_dStatusTelegramCounter := 1;
       ELSE
           #AUX_dStatusTelegramCounter += 1;
       END_IF;

       #ST_xStatusTelegramAvail := TRUE;

   END_IF;


   #AUX_xResetSendConnection := #IN_xGeneralReset OR (#FB_TSendSmall.s_TDIAG_Status.State <> b#16#04 AND #IN_xResetAlarms);


   IF (NOT #tPhasesNetworkSmall.xEndSendBuffer) AND (NOT #tPhasesNetworkSmall.xSendBuffer) AND 
           ((#ST_xRetrySendTelegramSmall)OR (#ST_xStatusTelegramAvail)OR (#ST_xDefectTelegramAvail) OR (#ST_xMessageTelegramAvail)) THEN

       IF (NOT #ST_xRetrySendTelegramSmall) THEN

           IF (#ST_xStatusTelegramAvail) THEN
               #TMP_dSerializePos := 0;
               #TMP_iReturn := Serialize(SRC_VARIABLE:=#AUX_tStatusPacket, DEST_ARRAY=>#AUX_rgb500SendBytePck, POS:=#TMP_dSerializePos);    
               #ST_xStatusTelegramAvail := FALSE;
           ELSIF (#ST_xDefectTelegramAvail) THEN
               #TMP_dSerializePos := 0;
               #TMP_iReturn := Serialize(SRC_VARIABLE:=#AUX_tDefectPacket, DEST_ARRAY=>#AUX_rgb500SendBytePck, POS:=#TMP_dSerializePos);    
               #ST_xDefectTelegramAvail := FALSE;
           ELSIF (#ST_xMessageTelegramAvail) THEN
               #TMP_dSerializePos := 0;
               #TMP_iReturn := Serialize(SRC_VARIABLE:=#AUX_tMessagePacketToOpt, DEST_ARRAY=>#AUX_rgb500SendBytePck, POS:=#TMP_dSerializePos);    
               #ST_xMessageTelegramAvail := FALSE;
           END_IF;

       END_IF;

       #ST_xRetrySendTelegramSmall := FALSE;
       #tPhasesNetworkSmall.xSendBuffer := TRUE;

   END_IF;

   #FB_TRecvSmall(EN_R:=TRUE,
                CONT:=TRUE,
                CONNECT:=#AUX_tConnDataSmall,
                DATA:=#AUX_rgb500RecvBytePck,
                COM_RST:=#AUX_xResetSendConnection);

   #FB_TRecvBig(EN_R:=TRUE,
                CONT:=TRUE,
               LEN := 0,
                CONNECT:=#AUX_tConnDataBig,
                DATA:=#AUX_rgb1000RecvBytePck,
                COM_RST:=#AUX_xResetSendConnection);

   #FB_TSendSmall(REQ:=#tPhasesNetworkSmall.xSendBuffer,
             CONT:=TRUE,
             LEN:=0,
             CONNECT:=#AUX_tConnDataSmall,
             DATA:=#AUX_rgb500SendBytePck,
             COM_RST:=#AUX_xResetSendConnection);

   #FB_TSendBig(REQ:=#tPhasesNetworkBig.xSendBuffer,
             CONT:=TRUE,
             LEN:=0,
             CONNECT:=#AUX_tConnDataBig,
             DATA:=#AUX_rgb1000SendBytePck,
             COM_RST:=#AUX_xResetSendConnection);

   //Manage send of the small packets
   IF #tPhasesNetworkSmall.xSendBuffer AND 
                                           (#FB_TSendSmall.DONE OR
                                           #FB_TSendSmall.ERROR OR 
                                           NOT #FB_TSendSmall.BUSY) THEN

       #tPhasesNetworkSmall.xSendBuffer := FALSE;
       #tPhasesNetworkSmall.xEndSendBuffer := TRUE;
       #ST_xRetrySendTelegramSmall := FALSE;

      IF NOT #FB_TSendSmall.DONE THEN

           #ST_xRetrySendTelegramSmall := TRUE;

       END_IF;



   ELSE

       #tPhasesNetworkSmall.xEndSendBuffer := FALSE;

   END_IF;

   //Manage received little telegram
   IF #FB_TRecvSmall.DONE THEN

       //Check the packet telegram
       #TMP_dSerializePos := 0;
       #TMP_iReturn := Deserialize(SRC_ARRAY:=#AUX_rgb500RecvBytePck, DEST_VARIABLE=>#TMP_dValue, POS:=#TMP_dSerializePos);

       IF #TMP_dValue = #DMESSAGERECVPACKETIDENT THEN

           #TMP_dSerializePos := 0;
           #TMP_iReturn := Deserialize(SRC_ARRAY:=#AUX_rgb500RecvBytePck, DEST_VARIABLE=>#AUX_tMessagePacketFromOpt, POS:=#TMP_dSerializePos);

           //Loop inside the packet and copy on the plc
           IF #AUX_tMessagePacketFromOpt.dNumMessage > 0 AND #AUX_tMessagePacketFromOpt.dNumMessage <= #DMAXMESSAGEPACKET THEN

               FOR #TMP_dIndex := 0 TO #AUX_tMessagePacketFromOpt.dNumMessage - 1 DO

                   "RP_AddMessageV2"(IN_xInit:=FALSE,
                                     IN_dCodeEvent:=#AUX_tMessagePacketFromOpt.rgtMessage[#TMP_dIndex].dCodeEvent,
                                     IN_strIndet_Max4Chars:='OPT',
                                     IN_dValue1:=#AUX_tMessagePacketFromOpt.rgtMessage[#TMP_dIndex].dEvent1,
                                     IN_dValue2:=#AUX_tMessagePacketFromOpt.rgtMessage[#TMP_dIndex].dEvent2,
                                     IN_dValue3:=#AUX_tMessagePacketFromOpt.rgtMessage[#TMP_dIndex].dEvent3,
                                     IN_dValue4:=#AUX_tMessagePacketFromOpt.rgtMessage[#TMP_dIndex].dEvent4,
                                     IN_dValue5:=#AUX_tMessagePacketFromOpt.rgtMessage[#TMP_dIndex].dEvent5,
                                     IN_dValue6:=#AUX_tMessagePacketFromOpt.rgtMessage[#TMP_dIndex].dEvent6,
                                     IN_dValue7:=#AUX_tMessagePacketFromOpt.rgtMessage[#TMP_dIndex].dEvent7,
                                     IN_dValue8:=#AUX_tMessagePacketFromOpt.rgtMessage[#TMP_dIndex].dEvent8,
                                     IN_dValue9:=#AUX_tMessagePacketFromOpt.rgtMessage[#TMP_dIndex].dEvent9,
                                     IN_dValue10:=#AUX_tMessagePacketFromOpt.rgtMessage[#TMP_dIndex].dEvent10,
                                     INO_tBuffer:=#INO_tAddMessageFromOpt,
                                     INO_xError:=#INO_xMessageAnomaly);

                   "RP_AddMessageV2"(IN_xInit:=FALSE,
                                     IN_dCodeEvent:=#AUX_tMessagePacketFromOpt.rgtMessage[#TMP_dIndex].dCodeEvent,
                                     IN_strIndet_Max4Chars:='OPT',
                                     IN_dValue1:=#AUX_tMessagePacketFromOpt.rgtMessage[#TMP_dIndex].dEvent1,
                                     IN_dValue2:=#AUX_tMessagePacketFromOpt.rgtMessage[#TMP_dIndex].dEvent2,
                                     IN_dValue3:=#AUX_tMessagePacketFromOpt.rgtMessage[#TMP_dIndex].dEvent3,
                                     IN_dValue4:=#AUX_tMessagePacketFromOpt.rgtMessage[#TMP_dIndex].dEvent4,
                                     IN_dValue5:=#AUX_tMessagePacketFromOpt.rgtMessage[#TMP_dIndex].dEvent5,
                                     IN_dValue6:=#AUX_tMessagePacketFromOpt.rgtMessage[#TMP_dIndex].dEvent6,
                                     IN_dValue7:=#AUX_tMessagePacketFromOpt.rgtMessage[#TMP_dIndex].dEvent7,
                                     IN_dValue8:=#AUX_tMessagePacketFromOpt.rgtMessage[#TMP_dIndex].dEvent8,
                                     IN_dValue9:=#AUX_tMessagePacketFromOpt.rgtMessage[#TMP_dIndex].dEvent9,
                                     IN_dValue10:=#AUX_tMessagePacketFromOpt.rgtMessage[#TMP_dIndex].dEvent10,
                                     INO_tBuffer:=#INO_tAddMessageToOpt,
                                     INO_xError:=#INO_xMessageAnomaly);

                   IF #AUX_tMessagePacketFromOpt.rgtMessage[#TMP_dIndex].dCodeEvent = "DEVENTS_MARKER_MISSION" THEN

                       #TMP_tNewMisMark.dMarkerID := #AUX_tMessagePacketFromOpt.rgtMessage[#TMP_dIndex].dEvent3;
                       #TMP_tNewMisMark.dMissionID := #AUX_tMessagePacketFromOpt.rgtMessage[#TMP_dIndex].dEvent2;
                       #TMP_tNewMisMark.dPlateID := #AUX_tMessagePacketFromOpt.rgtMessage[#TMP_dIndex].dEvent1;
                       #TMP_tNewMisMark.dSpotSpace_cmm := #AUX_tMessagePacketFromOpt.rgtMessage[#TMP_dIndex].dEvent6;
                       #TMP_tNewMisMark.dXPosition_cmm := #AUX_tMessagePacketFromOpt.rgtMessage[#TMP_dIndex].dEvent4;
                       #TMP_tNewMisMark.dYPosition_cmm := #AUX_tMessagePacketFromOpt.rgtMessage[#TMP_dIndex].dEvent5;
                       #TMP_xCallAddTank := TRUE;